(* Logix 5000 project; controller PLC_MCC1300_75F1 vendor 1 type 14 code 166 rev 32.11; software revision 32.04; part 59 of 83 *)
(* tags used below, declared in another part *)
   CONST_dDest_Cullet : DINT;
   CONST_dDest_Stk : DINT;
   CONST_rgdDestMask : DINT[32];   // Destination Mask
   GP_CheckIdPlatePresent : GP_CheckIdPlatePresent;
   GP_OB_InitializeMain : GP_OB_Initialize;
   GP_RampSpace : GP_RampSpace;
   GP_ScadaPlate : GP_ScadaPlate;
   Gp_SpaceConvUtilities_V1 : GP_SpaceConvUtilities_V1;
   M312 : MAC_Conveyor_Single;
   M312_ALM : MAC_Conveyor_ALM;
   M312_Data : UDT_Convoy_SL;
   M312_HMR : MAC_Conveyor_HMR;
   M312_SpaceConv_Utilities : SpaceConv_Utilities;
   M312_xLatLeftTimeout : BOOL;
   M315A : MAC_Conveyor;
   M315A_ALM : MAC_Conveyor_ALM;
   M315A_Data : UDT_Convoy_SL;
   M315A_dLastSyncID : DINT;
   M315A_HMR : MAC_Conveyor_HMR;
   M315A_HMW : MAC_Conveyor_HMW;
   M315A_INPUT_xSyncroPhotocell : BOOL;
   M315A_M1_DR : AXIS_CIP_DRIVE;
   M315A_OSR_xSyncOnLoad : BOOL;
   M315A_SpaceConv_Utilities : SpaceConv_Utilities;
   M315A_xSyncOnLoadDone : BOOL;
   M315B_SpaceConv_Utilities : SpaceConv_Utilities;
   M316 : MAC_Conveyor;
   M316_SpaceConv_Utilities : SpaceConv_Utilities;
   M317 : MAC_Conveyor_Single;
   M317_Data : UDT_Convoy_SL;
   O : INT[128];
   TMP_d : DINT;
   TMP_dConveyorNumberForZoneCleaning : DINT;
   TMP_dDecelerationPositionEndConveyor : DINT;
   TMP_dOffsetLoadUnload_cmm : DINT;
   TMP_rgxId : DINT[10];
   TMP_SendToCullet : BOOL;
   TMP_xConveyorInvolvedInCleaning : BOOL;
   TMP_xConveyorOfStartCleaning : BOOL;
   TMP_xCulletPresent : BOOL;
   TMP_xEnableLoadUnload : BOOL;
   TMP_xEnableZoneCleaning : BOOL;
   TMP_xLiteThisDestPresent : BOOL;
   xAlwaysOFF : BOOL;
   xAlwaysON : BOOL;
   Z401_HMI_rgtPlateScada_Internal : HMI_LiteData[5,2,7];
   Z402 : MAC_Zone;
   Z402_HMI_rgtPlateScada_Internal : HMI_LiteData[5,2,7];
   Z402_HMR : MAC_Zone_HMR;
   Z402_HMW : MAC_Zone_HMW;
(* MainProgram, continued *)

   // State Sensor
   123: XIC(xAlwaysON)[MOV(1,M312_HMR.dStateSensor2) ,[XIC(M312_ALM.rgxWarning[0].26) ,XIC(M312_xLatLeftTimeout) ] MOV(7,M312_HMR.dStateSensor2) ];
   124: XIC(M312.ST_xIdPlatePresence)GP_ScadaPlate(GP_ScadaPlate,M312_Data,6,M312_SpaceConv_Utilities.O_dHeadPosition_cmm,M312_SpaceConv_Utilities.CONST_dConveyorWidth_cmm,M312_SpaceConv_Utilities.CONST_dConveyorLength_cmm,M312_SpaceConv_Utilities.ST_xLastModLoadBkw,M312_SpaceConv_Utilities.ST_xLastModUnloadBkw,1,0,Z401_HMI_rgtPlateScada_Internal);
END_ROUTINE

ROUTINE M315A_Alarm   (* ladder *)
   // Reset Alarm
   0: XIC(Z402.tmON_ResetAlarm.DN)FLL(0,M315A_ALM,1);
   1: XIC(Z402.ST_xEnableControlError)XIC(xAlwaysOFF)XIO(M315A.INPUT_xProtectionMotor_M1)OTL(M315A_ALM.rgxStoppingFault_M[0].0);
   2: XIC(Z402.ST_xEnableControlError)XIC(M315A.INPUT_xDriveError_M1)OTL(M315A_ALM.rgxStoppingFault_M[0].1);
   3: XIC(Z402.ST_xEnableControlError)XIO(M315A.INPUT_xDriveError_M1)[XIC(M315A.OUTPUT_xRun_M1) ,XIC(M315A.OUTPUT_xReverse_M1) ,XIC(M315A.OUTPUT_xPositioning_M1) ]XIO(M315A.INPUT_xDriveFeedback_M1)[XIO(M315A.tmON_FeedbackTimeOut_M1.DN) TON(M315A.tmON_FeedbackTimeOut_M1,?,?) ,XIC(M315A.tmON_FeedbackTimeOut_M1.DN) OTL(M315A_ALM.rgxStoppingFault_M[0].2) ];
   4: XIC(Z402.ST_xEnableControlError)XIC(xAlwaysOFF)XIO(M315A.INPUT_xLocalSafetySwitch_M1)OTL(M315A_ALM.rgxStoppingFault_M[0].3);
   5: XIC(Z402.ST_xEnableControlError)XIO(M315A.INPUT_xMotorThermalProbe_M1)OTL(M315A_ALM.rgxStoppingFault_M[0].4);
   6: XIC(Z402.ST_xEnableControlError)XIC(xAlwaysOFF)XIO(M315A.INPUT_xBrakingResistor_M1)OTL(M315A_ALM.rgxStoppingFault_M[0].5);
   7: XIC(Z402.ST_xEnableControlError)[XIC(M315A.INPUT_xDriveInhibit_M1) ,XIC(M315A.OUTPUT_xDriveEnable_M1) XIO(M315A.INPUT_xDriveReady_M1) ][XIO(M315A.tmON_DriveInhibit_M1.DN) TON(M315A.tmON_DriveInhibit_M1,?,?) ,XIC(M315A.tmON_DriveInhibit_M1.DN) OTL(M315A_ALM.rgxStoppingFault_M[0].6) ];
   8: XIC(M315A.ST_xEnableControlError)XIC(M315A.PH_x.7)NEQ(M315A_SpaceConv_Utilities.CONST_dSyncMode,0)[XIO(M315A.ST_xPlateSynchronized) OTL(M315A_ALM.rgxWarning[0].0) ,XIC(M315A.ST_xPlateSynchronized) OTU(M315A_ALM.rgxWarning[0].0) ];
   9: XIC(M315A.ST_xEnableControlError)XIC(M315A.PH_x.7)[XIC(M315A_Data.tFlag.tConveyor.xReqStop) ,XIC(M315A_Data.tFlag.tConveyor.xBypassReqEndStop) ]OTL(M315A_ALM.rgxWarning[0].1);
   // #####_CUMULATIVE ALARM_#####
   10: NOP();
   11: [NEQ(M315A_ALM.rgxStoppingFault[0],0) ,NEQ(M315A_ALM.rgxStoppingFault_M[0],0) ,NEQ(M315A_ALM.rgxStoppingFault_M[1],0) ]OTE(M315A.ST_xStopMachineFault);
   12: [NEQ(M315A_ALM.rgxFault[0],0) ,NEQ(M315A_ALM.rgxFault_M[0],0) ,NEQ(M315A_ALM.rgxFault_M[1],0) ]OTE(M315A.ST_xStopNextCycleFault);
END_ROUTINE

ROUTINE M315A_Logic   (* ladder *)
   // #####_COSTANTS_#####
   0: [MOV(5010,TMP_dConveyorNumberForZoneCleaning) MOV(50000,TMP_dOffsetLoadUnload_cmm) MOV(500,M315A_SpaceConv_Utilities.CONST_dPresetFeedbackTime_ms) OTL(TMP_xEnableLoadUnload) OTL(TMP_xEnableZoneCleaning) MOV(800000,M315A_SpaceConv_Utilities.CONST_dConveyorLength_cmm) MOV(400000,M315A_SpaceConv_Utilities.CONST_dConveyorWidth_cmm) SUB(M315A_SpaceConv_Utilities.CONST_dConveyorLength_cmm,180000,M315A.AUX_dPresetStopLoad_cmm) ADD(M315A_SpaceConv_Utilities.CONST_dConveyorLength_cmm,M315A.AUX_dDecSpace_cmm,M315A.AUX_dPresetStopUnload_cmm) MOV(1.2,M315A_SpaceConv_Utilities.CONST_rAcceleration_ms2) MOV(1.2,M315A_SpaceConv_Utilities.CONST_rDeceleration_ms2) ,[MOV(1,M315A_SpaceConv_Utilities.CONST_dSyncMode) ,MOV(0,M315A_SpaceConv_Utilities.CONST_dSyncroPhPosition_cmm) ,MOV(450000,M315A_SpaceConv_Utilities.CONST_dSyncroPhWindow_cmm) ] ];
   // #####_MATCH_#####
   1: NOP();
   // Conveyor Cleaning
   2: XIC(TMP_xEnableZoneCleaning)XIC(Z402.ST_xCleaningAccepted)GRT(Z402_HMW.dCleaningSelection,0)[EQU(Z402_HMW.dCleaningSelection,TMP_dConveyorNumberForZoneCleaning) OTE(TMP_xConveyorOfStartCleaning) ,GEQ(Z402_HMW.dCleaningSelection,TMP_dConveyorNumberForZoneCleaning) OTE(TMP_xConveyorInvolvedInCleaning) ];
   // Enable control error
   3: XIC(Z402.ST_xEnableControlError)OTE(M315A.ST_xEnableControlError);
   // Mode 7 - Offsett for load/unload Simultaney
   4: XIC(M315A.PH_x.8)MOV(M315A.AUX_dPresetStopLoad_cmm,M315A_SpaceConv_Utilities.ST_dStopLoadForseen_cmm)MOV(TMP_dOffsetLoadUnload_cmm,M315A_SpaceConv_Utilities.CONF_MD7_dOffset_cmm)GP_SpaceConvUtilities_V1(Gp_SpaceConvUtilities_V1,M315A_SpaceConv_Utilities,M315B_SpaceConv_Utilities,M316_SpaceConv_Utilities,7);
   // #####_ALARMS_#####
   5: NOP();
   // Call Alarm Routine
   6: JSR(M315A_Alarm,0);
   // #####_HMI_LOGICS_#####
   7: NOP();
   // Condition ok for Cleaning
   8: [XIO(TMP_xEnableZoneCleaning) ,XIC(TMP_xEnableZoneCleaning) XIC(M315A.ST_xOutputEnable) [XIO(TMP_xConveyorOfStartCleaning) ,XIC(M315A.PH_x.0) ,XIO(M315A.PH_x.8) ] ]OTE(M315A.ST_xCleaningConditionOK);
   // Cleaning Accepted
   9: [[XIC(M315A_HMW.xStopLocalCleaningRequest) ,XIC(Z402_HMW.xStopCleanZoneRequest) ] OTU(M315A_HMW.xStopLocalCleaningRequest) OTU(M315A_HMW.xLocalCleaningRequest) ,[XIC(M315A_HMW.xLocalCleaningRequest) ,XIC(M317.ST_xCleaningAccepted) XIC(TMP_xEnableZoneCleaning) ] [XIC(M315A.ST_xCleaningConditionOK) ,XIC(M315A.ST_xCleaningAccepted) ] OTE(M315A.ST_xCleaningAccepted) ];
   // Manual Mode Enabled
   10: XIO(M315A_SpaceConv_Utilities.ST_xFeedbackRotation)[XIC(M315A_HMW.xEnableDisableManualCommand) XIC(M315A.ST_xConditionOKStopCycle) OTL(M315A.ST_xManualMode) ,XIO(M315A_HMW.xEnableDisableManualCommand) OTU(M315A.ST_xManualMode) ];
   // Virtual door enabled
   11: XIC(M315A_HMW.xEnableDisableVirtualDoor)OTE(M315A.ST_xVirtualDoorEnabled);
   // Clear manual command
   12: XIO(M315A.ST_xManualMode)MOV(0,M315A_HMW.rgxMan);
   // #####_STATUSES_#####
   13: NOP();
   // Syncro  -  OS Syncro Photocell
   14: XIC(xAlwaysON)[XIC(M315A_INPUT_xSyncroPhotocell) ONS(M315A.OSR_xSynchroPhotocellHead) OTE(M315A.OS_xSynchroPhotocellHead) GEQ(M315A_SpaceConv_Utilities.CONST_dSyncMode,1) OTE(M315A_SpaceConv_Utilities.ST_OS_xSynchroPhotocellHead) ,XIO(M315A_INPUT_xSyncroPhotocell) ONS(M315A.OSR_xSynchroPhotocellTail) OTE(M315A.OS_xSynchroPhotocellTail) GEQ(M315A_SpaceConv_Utilities.CONST_dSyncMode,2) OTE(M315A_SpaceConv_Utilities.ST_OS_xSynchroPhotocellTail) ];
   15: XIC(xAlwaysOFF)XIC(M315A_SpaceConv_Utilities.ST_OS_xSynchroPhotocellHead)XIO(M315A_xSyncOnLoadDone)ONS(M315A_OSR_xSyncOnLoad)XIC(M315A.PH_x.0)XIO(M315A.PH_x.8)GRT(M315A_Data.rgtCap[0].dID,0)NEQ(M315A_Data.rgtCap[0].dID,M315A_dLastSyncID)[MOV(0,M315A_SpaceConv_Utilities.CONF_MD2_MD3_dPrstPos_cmm) GP_SpaceConvUtilities_V1(Gp_SpaceConvUtilities_V1,M315A_SpaceConv_Utilities,M315B_SpaceConv_Utilities,M316_SpaceConv_Utilities,2) ,SUB(0,M315A_Data.dLength_cmm,M315A_SpaceConv_Utilities.CONF_MD2_MD3_dPrstPos_cmm) GP_SpaceConvUtilities_V1(Gp_SpaceConvUtilities_V1,M315A_SpaceConv_Utilities,M315B_SpaceConv_Utilities,M316_SpaceConv_Utilities,3) ,OTL(M315A_xSyncOnLoadDone) MOV(M315A_Data.rgtCap[0].dID,M315A_dLastSyncID) ];
   16: XIC(xAlwaysOFF)XIC(M315A.PH_x.0)XIC(M315A.OS_xSynchroPhotocellHead)XIO(M315A_xSyncOnLoadDone)[MOV(0,M315A_SpaceConv_Utilities.CONF_MD2_MD3_dPrstPos_cmm) GP_SpaceConvUtilities_V1(Gp_SpaceConvUtilities_V1,M315A_SpaceConv_Utilities,M315B_SpaceConv_Utilities,M316_SpaceConv_Utilities,2) ,SUB(0,M315A_Data.dLength_cmm,M315A_SpaceConv_Utilities.CONF_MD2_MD3_dPrstPos_cmm) GP_SpaceConvUtilities_V1(Gp_SpaceConvUtilities_V1,M315A_SpaceConv_Utilities,M315B_SpaceConv_Utilities,M316_SpaceConv_Utilities,3) ,OTL(M315A_xSyncOnLoadDone) ];
   // Id Plate presence
   17: MOV(CONST_rgdDestMask[24],CONST_dDest_Cullet)GP_CheckIdPlatePresent(GP_CheckIdPlatePresent,M315A_Data,TMP_rgxId,M315A.ST_xIdPlatePresence,TMP_xCulletPresent,CONST_dDest_Cullet)MOV(CONST_rgdDestMask[1],CONST_dDest_Stk)GP_CheckIdPlatePresent(GP_CheckIdPlatePresent,M315A_Data,TMP_rgxId,M315A.ST_xIdPlatePresence,TMP_xLiteThisDestPresent,CONST_dDest_Stk);
   // Machine in Alarm
   18: [XIC(M315A.ST_xStopMachineFault) ,XIC(M315A.ST_xStopNextCycleFault) ]OTE(M315A.ST_xMachineAlarm);
   // Condition ok for stop Cycle
   19: [XIO(M315A.ST_xPhasesInProgress) ,XIC(M315A.PH_x.8) XIO(M315A.OUTPUT_xRun_M1) XIO(M315A_SpaceConv_Utilities.ST_xFeedbackRotation) ,XIC(M315A.ST_xMachineAlarm) ,XIO(Z402.ST_xCycleON) ]OTE(M315A.ST_xConditionOKStopCycle);
   // Cycle load unload simultaneous
   20: XIC(TMP_xEnableLoadUnload)XIO(M315A.ST_xDisableLoadUnloadOnStop)XIO(M315A.ST_xIdPlatePresence)OTE(M315A.ST_xCycleLoadUnload);
   // Speed Management
   21: [XIO(M315A_SpaceConv_Utilities.O_xRampInProgress) XIO(M315A.ST_xManualMode) MOV(Z402_HMR.dLineSpeed_mm_min,M315A.AUX_dReqSpeed_mm_min) ,XIC(M315A.ST_xManualMode) MOV(Z402_HMW.dManualSpeed_mm_min,M315A.AUX_dReqSpeed_mm_min) ,NEQ(M315A.AUX_dReqSpeed_mm_min,M315A_SpaceConv_Utilities.ST_dRealSpeed_mm_min) OTE(M315A.OS_xChangeSpeed) ];
   // Ramp Management
   22: GP_RampSpace(GP_RampSpace,M315A_SpaceConv_Utilities.CONST_rAcceleration_ms2,M315A_SpaceConv_Utilities.CONST_rDeceleration_ms2,M315A_SpaceConv_Utilities.ST_dRealSpeed_mm_min,M315A.AUX_dAccSpace_cmm,M315A.AUX_dDecSpace_cmm);
   // Space Convoy utilities MOD 1 for Calculate Head/Tail
   23: XIC(xAlwaysON)[[XIC(M315A.OUTPUT_xRun_M1) ,XIC(M315A.OUTPUT_xReverse_M1) ] [XIO(M315A.ST_xManualMode) ,XIO(xAlwaysOFF) ] OTE(M315A_SpaceConv_Utilities.CONF_MD1_xRun) ,XIC(M315A.OUTPUT_xReverse_M1) XIC(xAlwaysOFF) XIO(M315A.ST_xManualMode) OTE(M315A_SpaceConv_Utilities.CONF_MD1_xReverse) ,[XIC(M315A.INPUT_xDriveFeedback_M1) ,XIC(M315A_SpaceConv_Utilities.CONF_MD1_xRun) GRT(M315A_SpaceConv_Utilities.O_dCountFeedbackTime_ms,0) ] OTE(M315A_SpaceConv_Utilities.ST_xFeedbackRotation) ,XIC(M315A.ST_xIdPlatePresence) OTE(M315A_SpaceConv_Utilities.CONF_MD1_xHeadTracking) ,XIC(M315A.ST_xPlatePresence) OTE(M315A_SpaceConv_Utilities.CONF_MD1_xTailTracking) ,MOV(GP_OB_InitializeMain.OUT_dExecutionTime_ms,M315A_SpaceConv_Utilities.CONF_MD1_dScan_ms) GP_SpaceConvUtilities_V1(Gp_SpaceConvUtilities_V1,M315A_SpaceConv_Utilities,M315B_SpaceConv_Utilities,M316_SpaceConv_Utilities,1) ];
   // Output Enable
   24: XIC(Z402.ST_xCycleON)XIO(M315A.ST_xManualMode)XIO(M315A.ST_xStopMachineFault)[XIO(M315A.ST_xPlatePassageUpstream_FW) XIO(M315A.ST_xPlatePassageUpstream_BKW) ,XIC(M315A.ST_xPlatePassageUpstream_FW) XIC(M317.ST_xOutputEnable) ]OTE(M315A.ST_xOutputEnable);
   // #####_WORKING_FLAGS_#####
   25: NOP();
   // #####_LOGICS_#####
   26: NOP();
   // Phase of load
   27: XIC(M317.OS_xUnload_FW)[OTL(M315A.PH_x.0) ,OTU(M315A_SpaceConv_Utilities.O_xPlateSynchronized) ,OTU(M315A.ST_xDisableLoadUnloadOnStop) ,OTE(M315A.OS_xLoad_FW) ,COP(M317_Data,M315A_Data,1) FLL(0,M317_Data,1) ,GP_SpaceConvUtilities_V1(Gp_SpaceConvUtilities_V1,M315A_SpaceConv_Utilities,M315B_SpaceConv_Utilities,M316_SpaceConv_Utilities,5) ];
   // Syncro  -  Space Convoy utilities MOD 4
   28: GRT(M315A_SpaceConv_Utilities.CONST_dSyncMode,0)[XIC(M315A.PH_x.0) XIO(M315A.PH_x.8) ,XIC(M315A.PH_x.0) XIC(M315A.PH_x.8) ADD(M315A_SpaceConv_Utilities.CONST_dSyncroPhPosition_cmm,TMP_dOffsetLoadUnload_cmm,TMP_d) GRT(M315A_SpaceConv_Utilities.O_dTailPosition_cmm,TMP_d) ][MOV(M315A_Data.dLength_cmm,M315A_SpaceConv_Utilities.CONF_MD4_MD6_dLength_cmm) ,GP_SpaceConvUtilities_V1(Gp_SpaceConvUtilities_V1,M315A_SpaceConv_Utilities,M315B_SpaceConv_Utilities,M316_SpaceConv_Utilities,4) ];
   // End load Phase
   29: XIC(M315A.PH_x.0)GRT(M315A_SpaceConv_Utilities.O_dHeadPosition_cmm,M315A.AUX_dPresetStopLoad_cmm)[OTE(M315A.PH_x.7) ,OTU(M315A.PH_x.0) ,OTL(M315A.ST_xPlatePresence) ,OTU(M315A_xSyncOnLoadDone) ];
   // Calculation Space for Wait Stop Next Conveyor
   30: CPT(TMP_dDecelerationPositionEndConveyor,M315A_SpaceConv_Utilities.CONST_dConveyorLength_cmm - M315A.AUX_dAccSpace_cmm + 1000);
   // Wait stop next Machine
   31: XIO(M315A.PH_x.8)GEQ(M315A_SpaceConv_Utilities.O_dHeadPosition_cmm,TMP_dDecelerationPositionEndConveyor)OTE(M315A.ST_xWaitStopNextMachine);
   // Set Wait Machine Stop
   32: [XIC(M315A.PH_x.7) [XIO(M316.ST_xInitialConditionOK) ,XIC(M315A.ST_xWaitStopNextMachine) [XIC(M316_SpaceConv_Utilities.O_xRampInProgress) ,XIO(M316_SpaceConv_Utilities.ST_xFeedbackRotation) ] ] ,XIC(M315A.PH_x.0) NEQ(Z402_HMR.dLineSpeed_mm_min,M315A.AUX_dReqSpeed_mm_min) ]OTL(M315A.ST_xWaitMachineStop);
   // Reset Wait Machine Stop
   33: XIO(M315A_SpaceConv_Utilities.ST_xFeedbackRotation)[XIO(M315A_SpaceConv_Utilities.ST_xFeedbackRotation) ,XIO(M315A.ST_xWaitStopNextMachine) ]EQU(Z402_HMR.dLineSpeed_mm_min,M315A.AUX_dReqSpeed_mm_min)OTU(M315A.ST_xWaitMachineStop);
   // Phase of unload
   34: XIC(Z402.ST_xConditionOkPhaseAdvancement)XIC(M315A.ST_xPlatePresence)XIC(M315A.ST_xIdPlatePresence)XIC(M315A.ST_xOutputEnable)XIC(M316.ST_xInitialConditionOK)XIO(M315A.ST_xWaitMachineStop)XIO(M315A.PH_x.8)[OTE(M315A.ST_xWaitReadyToMove) ,[XIC(M315A.ST_xAxleReadyToMoveDelayed) ,XIC(xAlwaysON) ] [OTE(M315A.OS_xUnload_FW) ,OTL(M315A.PH_x.8) ,MOV(M315A_Data.dLength_cmm,M315A_SpaceConv_Utilities.CONF_MD4_MD6_dLength_cmm) GP_SpaceConvUtilities_V1(Gp_SpaceConvUtilities_V1,M315A_SpaceConv_Utilities,M315B_SpaceConv_Utilities,M316_SpaceConv_Utilities,6) ] ];
   // Phase of end unload
   35: XIC(M315A.PH_x.8)[GEQ(M315A_SpaceConv_Utilities.O_dTailPosition_cmm,M315A.AUX_dPresetStopUnload_cmm) ,XIO(M315A_SpaceConv_Utilities.ST_xFeedbackRotation) GEQ(M315A_SpaceConv_Utilities.O_dTailPosition_cmm,M315A_SpaceConv_Utilities.CONST_dConveyorLength_cmm) ][OTE(M315A.PH_x.15) ,OTU(M315A.PH_x.8) ,OTU(M315A.ST_xPlatePresence) ];
   // Phase in progress
   36: NEQ(M315A.PH_x,0)OTE(M315A.ST_xPhasesInProgress);
   // #####_CLEANING_#####
   37: NOP();
   // Cleaning Reset
   38: XIC(M315A.ST_xCleaningAccepted)[XIC(Z402.ST_xCleaningAccepted) ,XIO(TMP_xConveyorOfStartCleaning) ][XIC(M315A.ST_xIdPlatePresence) OTL(TMP_SendToCullet) FLL(0,M315A_Data,1) ,MOV(0,M315A.PH_x) OTU(M315A.ST_xPlatePresence) ];
   // Initial condition OK
   39: XIC(Z402.ST_xConditionOkPhaseAdvancement)XIC(M315A.ST_xOutputEnable)XIO(M315A_HMW.xEnableDisableManualCommand)XIO(M315A.ST_xReqCleaning)XIO(M315A.ST_xCleaningAccepted)XIO(M315A.ST_xStopNextCycleFault)XIO(M315A.ST_xVirtualDoorEnabled)XIO(M315A.PH_x.0)[XIO(M315A.ST_xPhasesInProgress) XIO(M315A.ST_xPlatePresence) ,XIC(M315A.ST_xCycleLoadUnload) XIC(M315A.PH_x.8) XIC(M315A.OUTPUT_xRun_M1) GRT(M315A_SpaceConv_Utilities.O_dTailPosition_cmm,M315A_SpaceConv_Utilities.O_dPresetLoadUnload_cmm) XIO(M315A.ST_xIdPlatePresence) ]OTE(M315A.ST_xInitialConditionOK);
   // #####_HMI_STATUSES_#####
   40: NOP();
   // PhotocelPresence {x|x|x|x|O}
   41: XIC(M315A_INPUT_xSyncroPhotocell)OTE(M315A_HMR.xSensorPresence1);
   // Manual Mode Enable {x|x|x|x|O}
   42: XIC(M315A.ST_xManualMode)OTE(M315A_HMR.xManualCommandEnabled);
   // Command forward M1
   43: XIC(M315A.ST_xManualMode)XIC(M315A_HMW.rgxMan.0)XIC(M315A.OUTPUT_xRun_M1)OTE(M315A_HMR.rgxMan.0);
   // Command backward M1
   44: XIC(M315A.ST_xManualMode)XIC(M315A_HMW.rgxMan.1)XIC(M315A.OUTPUT_xReverse_M1)OTE(M315A_HMR.rgxMan.1);
   // Cleaning Enabled {x|x|x|x|O}
   45: XIC(M315A.ST_xCleaningAccepted)[XIC(Z402.ST_xCleaningAccepted) ,XIO(TMP_xEnableZoneCleaning) ]OTE(M315A_HMR.xCleaningEnabled);
   // Virtual door Enabled {x|x|x|x|O}
   46: XIC(M315A.ST_xVirtualDoorEnabled)OTE(M315A_HMR.xVirtualDoorEnabled);
   // Id plate presence
   47: XIC(M315A.ST_xIdPlatePresence)OTE(M315A_HMR.xIdPlatePresence);
   // Machine state M1
   48: XIC(xAlwaysON)[MOV(1,M315A_HMR.dState1) ,XIC(M315A.OUTPUT_xRun_M1) MOV(3,M315A_HMR.dState1) ,XIC(M315A.OUTPUT_xReverse_M1) MOV(4,M315A_HMR.dState1) ,XIC(M315A.ST_xMachineAlarm) MOV(7,M315A_HMR.dState1) ];
   49: XIC(M315A_SpaceConv_Utilities.O_xPlateSynchronized)OTE(M315A.ST_xPlateSynchronized);
   // State Sensor
   50: XIC(xAlwaysON)[MOV(1,M315A_HMR.dStateSensor1) ,XIC(M315A_ALM.rgxWarning[0].0) MOV(7,M315A_HMR.dStateSensor1) ];
   // Motor error code
   51: MOV(M315A_M1_DR.AxisFault,M315A_HMR.dErrorCode1);
   52: XIC(M315A.ST_xIdPlatePresence)GP_ScadaPlate(GP_ScadaPlate,M315A_Data,1,M315A_SpaceConv_Utilities.O_dHeadPosition_cmm,M315A_SpaceConv_Utilities.CONST_dConveyorWidth_cmm,M315A_SpaceConv_Utilities.CONST_dConveyorLength_cmm,0,0,1,1,Z402_HMI_rgtPlateScada_Internal);
END_ROUTINE
